// TIA Portal project "DATN" (V16)

(* hardware
DEVICE "S7-1200 station_1"  S7-1200 Station
   slot 0: "Rack_0"  S7-1200 Rack  Rack  V1.0
   slot 1: "PLC_1"  CPU 1214C DC/DC/DC  6ES7 214-1AG40-0XB0  V4.0
DEVICE "PC-System_1"  SIMATIC PC station
   slot 0: "SIMATIC PC station"  Rail  SIMATIC PC-Station  V1.0
      slot 125: "Stationmanager"  Station_Manager  V6.0.4
   slot 1: "HMI_RT_1"  WinCC RT Advanced  6AV2 104-0xxxx-xxxx  16.0.0.0
      slot 33792: "Computer interface"  Host interface
   slot 2: "IE general_1"  IE General  IE_CP  V8.2.0
*)

// ===== PLC "PLC_1"  CPU 1214C DC/DC/DC =====

VAR_GLOBAL   // PLC tag table "Default tag table"
   "System_Byte" AT %MB1000 : Byte;
   "FirstScan" AT %M1000.0 : Bool;
   "DiagStatusUpdate" AT %M1000.1 : Bool;
   "AlwaysTRUE" AT %M1000.2 : Bool;
   "AlwaysFALSE" AT %M1000.3 : Bool;
END_VAR

VAR_GLOBAL   // PLC tag table "1_IN"
   "CB_CAP_PHOI" AT %I0.0 : Bool;
   "CB_SP_1" AT %I0.1 : Bool;
   "CB_SP_2" AT %I0.2 : Bool;
   "CB_SP_3" AT %I0.3 : Bool;
   "PB_START" AT %I0.4 : Bool;
   "PB_STOP" AT %I0.5 : Bool;
   "PB_RESET" AT %I0.6 : Bool;
   "HMI_CB_CAP_PHOI" AT %M100.0 : Bool;
   "HMI_CB_SP_1" AT %M100.1 : Bool;
   "HMI_CB_SP_2" AT %M100.2 : Bool;
   "HMI_CB_SP_3" AT %M100.3 : Bool;
   "HMI_PB_START" AT %M100.4 : Bool;
   "HMI_PB_STOP" AT %M100.5 : Bool;
   "HMI_PB_RESET" AT %M100.6 : Bool;
   "MAN_BT" AT %M100.7 : Bool;
   "MAN_XYLANH_1" AT %M101.0 : Bool;
   "MAN_XYLANH_2" AT %M101.1 : Bool;
   "MAN_CAP_PHOI" AT %M101.2 : Bool;
   "HMI_AUTO_MAN" AT %M101.3 : Bool;
   "RST_SP_1" AT %M101.4 : Bool;
   "RST_SP_2" AT %M101.5 : Bool;
   "RST_SP_3" AT %M101.6 : Bool;
END_VAR

VAR_GLOBAL   // PLC tag table "2_OUT"
   "BANG_TAI" AT %Q0.0 : Bool;
   "XY_LANH_1" AT %Q0.1 : Bool;
   "XY_LANH_2" AT %Q0.2 : Bool;
   "DEN_START" AT %Q0.5 : Bool;
   "DEN_STOP" AT %Q0.6 : Bool;
   "XY_LANH_CAP_PHOI_1" AT %Q0.3 : Bool;
   "DEN_RESET" AT %Q0.7 : Bool;
END_VAR

VAR_GLOBAL   // PLC tag table "3_MEMORY"
   "SP_3" AT %M200.0 : Bool;
   "RUN_PHAN_LOAI" AT %M200.1 : Bool;
   "BT_1" AT %M200.2 : Bool;
   "BT_2" AT %M200.3 : Bool;
   "NGAT_CB_CAP_PHOI" AT %M200.4 : Bool;
   "RST_COUNTER_SP_1" AT %M200.5 : Bool;
   "RST_COUNTER_SP_2" AT %M200.6 : Bool;
   "RST_COUNTER_SP_3" AT %M200.7 : Bool;
   "den_rst_1" AT %M201.1 : Bool;
   "den_rst_2" AT %M201.2 : Bool;
   "NGAT_HE_THONG" AT %M201.3 : Bool;
   "OUT_counter_1" AT %M201.4 : Bool;
   "OUT_counter_2" AT %M201.5 : Bool;
   "OUT_counter_3" AT %M201.6 : Bool;
   "MODE_AUTO" AT %M201.7 : Bool;
   "MODE_MAN" AT %M202.0 : Bool;
   "xylanh_cap_phoi_auto" AT %M202.1 : Bool;
   "xylanh_cap_phoi_man" AT %M202.2 : Bool;
   "xylanh_1_auto" AT %M202.3 : Bool;
   "xylanh_1_man" AT %M202.4 : Bool;
   "xylanh_2_auto" AT %M202.5 : Bool;
   "xylanh_2_man" AT %M202.6 : Bool;
   "ngat_mau_sac" AT %M202.7 : Bool;
END_VAR

VAR_GLOBAL   // PLC tag table "5_M_TIME_500"
   "TIME_XY_LANH_1" AT %MD500 : Time;
   "TIME_XY_LANH_2" AT %MD504 : Time;
   "TIME_SP_3" AT %MD508 : Time;
   "TIME_CAP_PHOI" AT %MD512 : Time;
   "TIME_NGAT_CAP_PHOI" AT %MD516 : Time;
   "TIME_ERROR_KHONG_SP" AT %MD520 : Time;
   "TIME_ERROR_STUCK" AT %MD524 : Time;
END_VAR

VAR_GLOBAL   // PLC tag table "4_P_N_MEMORy"
   "N_CB_SP_1" AT %M300.0 : Bool;
   "N_CB_SP_2" AT %M300.1 : Bool;
   "N_CB_SP_3" AT %M300.2 : Bool;
   "N_XY_LANH_1" AT %M300.3 : Bool;
   "N_XY_LANH_2" AT %M300.4 : Bool;
   "N_SP_3" AT %M300.5 : Bool;
   "N_M_CB_SP_1" AT %M300.6 : Bool;
   "N_M_CB_SP_2" AT %M300.7 : Bool;
   "N_M_CB_SP_3" AT %M301.0 : Bool;
END_VAR

VAR_GLOBAL   // PLC tag table "6_DATA_real_int"
   "LUU_MAU" AT %MW222 : Int;
   "Mau Sac" AT %MW220 : Int;
END_VAR

VAR_GLOBAL   // PLC tag table "7_ALARM"
   "BIT_WARNING_KHONG_SP" AT %M400.0 : Bool;
   "DATA_WORD_WARNING" AT %MW400 : Int;
   "MULTI_ERROR" AT %M450.0 : Bool;
   "BIT_ERROR_STUCK_sp_1" AT %M402.0 : Bool;
   "BIT_ERROR_STUCK_sp_2" AT %M404.0 : Bool;
   "BIT_ERROR_STUCK_sp_3" AT %M406.0 : Bool;
   "DATA_WORD_ERROR_1" AT %MW402 : Int;
   "DATA_WORD_ERROR_2" AT %MW404 : Int;
   "DATA_WORD_ERROR_3" AT %MW406 : Int;
END_VAR

DATA_BLOCK "MB"   // DB12
{ S7_Optimized_Access := 'FALSE' }
VERSION : 0.1
   VAR
      DISCONNECT : Bool;
      H_reg : Array[0..10] of Int;
      CONNECT : TCON_IP_v4;
      ERROR : Bool;
      STATUS : Word;
   END_VAR
BEGIN
   CONNECT.InterfaceId := 64;
   CONNECT.ID := 1;
   CONNECT.ConnectionType := 11;
   CONNECT.ActiveEstablished := TRUE;
   CONNECT.RemoteAddress.ADDR[1] := 192;
   CONNECT.RemoteAddress.ADDR[2] := 168;
   CONNECT.RemoteAddress.ADDR[3] := 0;
   CONNECT.RemoteAddress.ADDR[4] := 10;
   CONNECT.LocalPort := 502;
   CONNECT.RemotePort := 0;
END_DATA_BLOCK

DATA_BLOCK "gh_sp"   // DB13
{ S7_Optimized_Access := 'TRUE' }
VERSION : 0.1
   VAR
      GH_SP_1 : USInt := 3;
      GH_SP_2 : USInt := 3;
      GH_SP_3 : USInt := 3;
   END_VAR
BEGIN
END_DATA_BLOCK

// folder: System blocks/Program resources

DATA_BLOCK "TIMER_CAP_PHOI"   // DB1
{ S7_Optimized_Access := 'TRUE' }
AUTHOR : Simatic
FAMILY : IEC
NAME : IEC_TMR
VERSION : 1.0
// stored: InstanceOfName IEC_TIMER
"IEC_TIMER"
BEGIN
END_DATA_BLOCK

DATA_BLOCK "TIMER_XY_LANH_1"   // DB2
{ S7_Optimized_Access := 'TRUE' }
AUTHOR : Simatic
FAMILY : IEC
NAME : IEC_TMR
VERSION : 1.0
// stored: InstanceOfName IEC_TIMER
"IEC_TIMER"
BEGIN
END_DATA_BLOCK

DATA_BLOCK "TIMER_XY_LANH_2"   // DB3
{ S7_Optimized_Access := 'TRUE' }
AUTHOR : Simatic
FAMILY : IEC
NAME : IEC_TMR
VERSION : 1.0
// stored: InstanceOfName IEC_TIMER
"IEC_TIMER"
BEGIN
END_DATA_BLOCK

DATA_BLOCK "TIMER_SP_3"   // DB4
{ S7_Optimized_Access := 'TRUE' }
AUTHOR : Simatic
FAMILY : IEC
NAME : IEC_TMR
VERSION : 1.0
// stored: InstanceOfName IEC_TIMER
"IEC_TIMER"
BEGIN
END_DATA_BLOCK

DATA_BLOCK "COUNTER_SP_1"   // DB5
{ S7_Optimized_Access := 'TRUE' }
AUTHOR : Simatic
FAMILY : IEC
NAME : CNTR
VERSION : 1.0
// stored: InstanceOfName IEC_COUNTER
"IEC_COUNTER"
BEGIN
END_DATA_BLOCK

DATA_BLOCK "COUNTER_SP_2"   // DB6
{ S7_Optimized_Access := 'TRUE' }
AUTHOR : Simatic
FAMILY : IEC
NAME : CNTR
VERSION : 1.0
// stored: InstanceOfName IEC_COUNTER
"IEC_COUNTER"
BEGIN
END_DATA_BLOCK

DATA_BLOCK "COUNTER_SP_3"   // DB7
{ S7_Optimized_Access := 'TRUE' }
AUTHOR : Simatic
FAMILY : IEC
NAME : CNTR
VERSION : 1.0
// stored: InstanceOfName IEC_COUNTER
"IEC_COUNTER"
BEGIN
END_DATA_BLOCK

DATA_BLOCK "TIMER_NGAT_CAP_PHOI"   // DB8
{ S7_Optimized_Access := 'TRUE' }
AUTHOR : Simatic
FAMILY : IEC
NAME : IEC_TMR
VERSION : 1.0
// stored: InstanceOfName IEC_TIMER
"IEC_TIMER"
BEGIN
END_DATA_BLOCK

DATA_BLOCK "TIMER_LOI_KHONG_SP"   // DB9
{ S7_Optimized_Access := 'TRUE' }
AUTHOR : Simatic
FAMILY : IEC
NAME : IEC_TMR
VERSION : 1.0
// stored: InstanceOfName IEC_TIMER
"IEC_TIMER"
BEGIN
END_DATA_BLOCK

DATA_BLOCK "TIMER_den_vang"   // DB10
{ S7_Optimized_Access := 'TRUE' }
AUTHOR : Simatic
FAMILY : IEC
NAME : IEC_TMR
VERSION : 1.0
// stored: InstanceOfName IEC_TIMER
"IEC_TIMER"
BEGIN
END_DATA_BLOCK

DATA_BLOCK "TIMER_STUCK_1"   // DB14
{ S7_Optimized_Access := 'TRUE' }
AUTHOR : Simatic
FAMILY : IEC
NAME : IEC_TMR
VERSION : 1.0
// stored: InstanceOfName IEC_TIMER
"IEC_TIMER"
BEGIN
END_DATA_BLOCK

DATA_BLOCK "TIMER_STUCK_2"   // DB15
{ S7_Optimized_Access := 'TRUE' }
AUTHOR : Simatic
FAMILY : IEC
NAME : IEC_TMR
VERSION : 1.0
// stored: InstanceOfName IEC_TIMER
"IEC_TIMER"
BEGIN
END_DATA_BLOCK

DATA_BLOCK "TIMER_STUCK_3"   // DB16
{ S7_Optimized_Access := 'TRUE' }
AUTHOR : Simatic
FAMILY : IEC
NAME : IEC_TMR
VERSION : 1.0
// stored: InstanceOfName IEC_TIMER
"IEC_TIMER"
BEGIN
END_DATA_BLOCK

// folder: (top level)

FUNCTION "FC_1_Modbus_TCP" : Void   // FC1, LAD
{ S7_Optimized_Access := 'TRUE' }
VERSION : 0.1
BEGIN

REGION Network 1
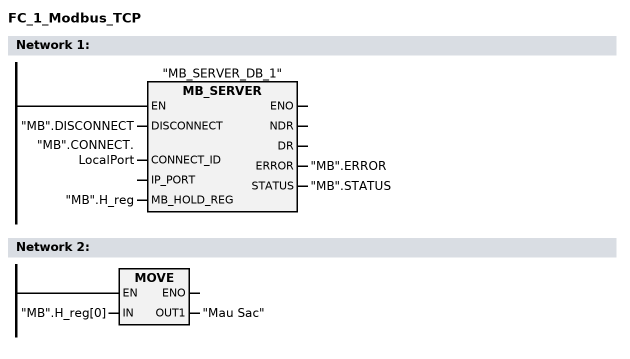
   "MB_SERVER_DB_1"(DISCONNECT := "MB".DISCONNECT,   // MB_SERVER
                    CONNECT_ID := "MB".CONNECT.LocalPort,
                    MB_HOLD_REG := "MB".H_reg,
                    ERROR => "MB".ERROR,
                    STATUS => "MB".STATUS);
END_REGION

REGION Network 2
   RUNG wire#powerrail
      Move(in := "MB".H_reg[0], out1 => "Mau Sac")
   END_RUNG
   // the same network as SCL:
   "Mau Sac" := "MB".H_reg[0];
END_REGION
END_FUNCTION

FUNCTION "FC_4_PHAN_LOAI_SP_1" : Void   // FC2, LAD
{ S7_Optimized_Access := 'TRUE' }
VERSION : 0.1
   VAR_TEMP   // added for the SCL form of the ladder/FBD networks
      _w1 : Bool;
      _w2 : Bool;
   END_VAR
BEGIN

REGION Network 1
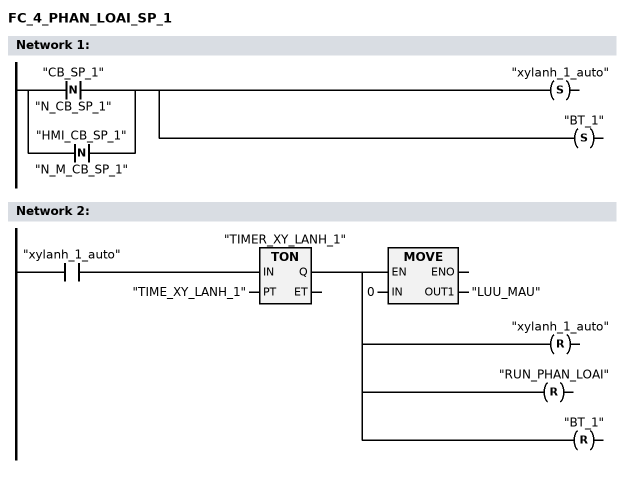
   RUNG wire#powerrail
      N_Contact(operand := "CB_SP_1", bit := "N_CB_SP_1")
      wire#w1
      S_Coil( "xylanh_1_auto" )
   END_RUNG
   RUNG wire#powerrail
      N_Contact(operand := "HMI_CB_SP_1", bit := "N_M_CB_SP_1")
   END_RUNG wire#w1
   RUNG wire#w1
      S_Coil( "BT_1" )
   END_RUNG
   // the same network as SCL:
   #_w1 := NOT "CB_SP_1" AND "N_CB_SP_1";   // falling edge of "CB_SP_1"
   "N_CB_SP_1" := "CB_SP_1";
   #_w2 := NOT "HMI_CB_SP_1" AND "N_M_CB_SP_1";   // falling edge of "HMI_CB_SP_1"
   "N_M_CB_SP_1" := "HMI_CB_SP_1";
   IF #_w1 OR #_w2 THEN
       "xylanh_1_auto" := TRUE;
       "BT_1" := TRUE;
   END_IF;
END_REGION

REGION Network 2
   "TIMER_XY_LANH_1".TON(IN := "xylanh_1_auto", PT := "TIME_XY_LANH_1");
   IF "TIMER_XY_LANH_1".Q THEN
       "LUU_MAU" := 0;
       "xylanh_1_auto" := FALSE;
       "RUN_PHAN_LOAI" := FALSE;
       "BT_1" := FALSE;
   END_IF;
END_REGION
END_FUNCTION

FUNCTION "FC_5_PHAN_LOAI_SP_2" : Void   // FC3, LAD
{ S7_Optimized_Access := 'TRUE' }
VERSION : 0.1
   VAR_TEMP   // added for the SCL form of the ladder/FBD networks
      _w1 : Bool;
      _w2 : Bool;
   END_VAR
BEGIN

REGION Network 1
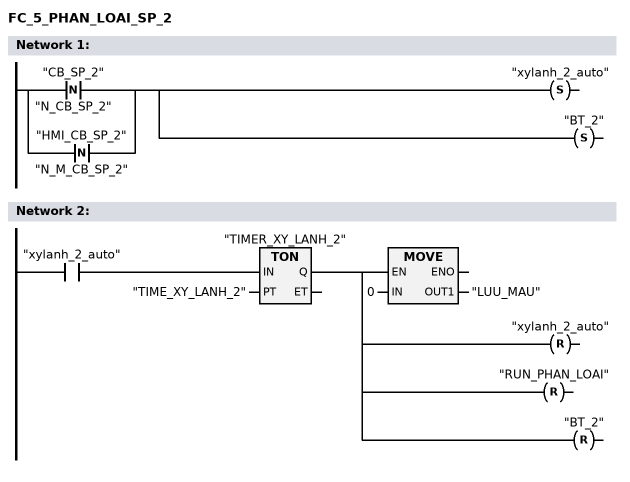
   RUNG wire#powerrail
      N_Contact(operand := "CB_SP_2", bit := "N_CB_SP_2")
      wire#w1
      S_Coil( "xylanh_2_auto" )
   END_RUNG
   RUNG wire#powerrail
      N_Contact(operand := "HMI_CB_SP_2", bit := "N_M_CB_SP_2")
   END_RUNG wire#w1
   RUNG wire#w1
      S_Coil( "BT_2" )
   END_RUNG
   // the same network as SCL:
   #_w1 := NOT "CB_SP_2" AND "N_CB_SP_2";   // falling edge of "CB_SP_2"
   "N_CB_SP_2" := "CB_SP_2";
   #_w2 := NOT "HMI_CB_SP_2" AND "N_M_CB_SP_2";   // falling edge of "HMI_CB_SP_2"
   "N_M_CB_SP_2" := "HMI_CB_SP_2";
   IF #_w1 OR #_w2 THEN
       "xylanh_2_auto" := TRUE;
       "BT_2" := TRUE;
   END_IF;
END_REGION

REGION Network 2
   "TIMER_XY_LANH_2".TON(IN := "xylanh_2_auto", PT := "TIME_XY_LANH_2");
   IF "TIMER_XY_LANH_2".Q THEN
       "LUU_MAU" := 0;
       "xylanh_2_auto" := FALSE;
       "RUN_PHAN_LOAI" := FALSE;
       "BT_2" := FALSE;
   END_IF;
END_REGION
END_FUNCTION

FUNCTION "FC_6_PHAN_LOAI_SP_3" : Void   // FC4, LAD
{ S7_Optimized_Access := 'TRUE' }
VERSION : 0.1
   VAR_TEMP   // added for the SCL form of the ladder/FBD networks
      _w1 : Bool;
      _w2 : Bool;
   END_VAR
BEGIN

REGION Network 1
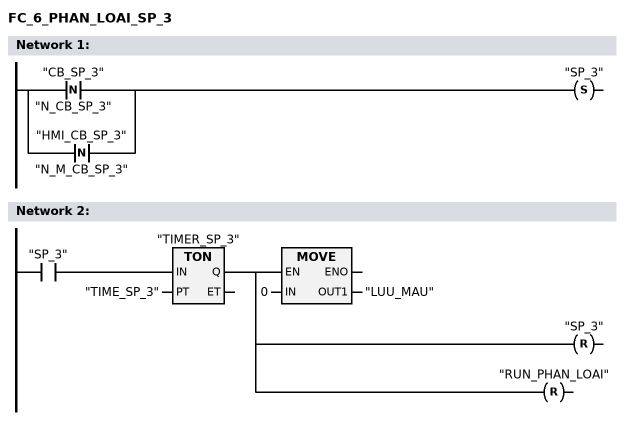
   RUNG wire#powerrail
      N_Contact(operand := "CB_SP_3", bit := "N_CB_SP_3")
      wire#w1
      S_Coil( "SP_3" )
   END_RUNG
   RUNG wire#powerrail
      N_Contact(operand := "HMI_CB_SP_3", bit := "N_M_CB_SP_3")
   END_RUNG wire#w1
   // the same network as SCL:
   #_w1 := NOT "CB_SP_3" AND "N_CB_SP_3";   // falling edge of "CB_SP_3"
   "N_CB_SP_3" := "CB_SP_3";
   #_w2 := NOT "HMI_CB_SP_3" AND "N_M_CB_SP_3";   // falling edge of "HMI_CB_SP_3"
   "N_M_CB_SP_3" := "HMI_CB_SP_3";
   IF #_w1 OR #_w2 THEN "SP_3" := TRUE; END_IF;
END_REGION

REGION Network 2
   "TIMER_SP_3".TON(IN := "SP_3", PT := "TIME_SP_3");
   IF "TIMER_SP_3".Q THEN
       "LUU_MAU" := 0;
       "SP_3" := FALSE;
       "RUN_PHAN_LOAI" := FALSE;
   END_IF;
END_REGION
END_FUNCTION

FUNCTION "FC_3_CAP_PHOI_TU_DONG" : Void   // FC5, LAD
{ S7_Optimized_Access := 'TRUE' }
VERSION : 0.1
BEGIN

REGION Network 1
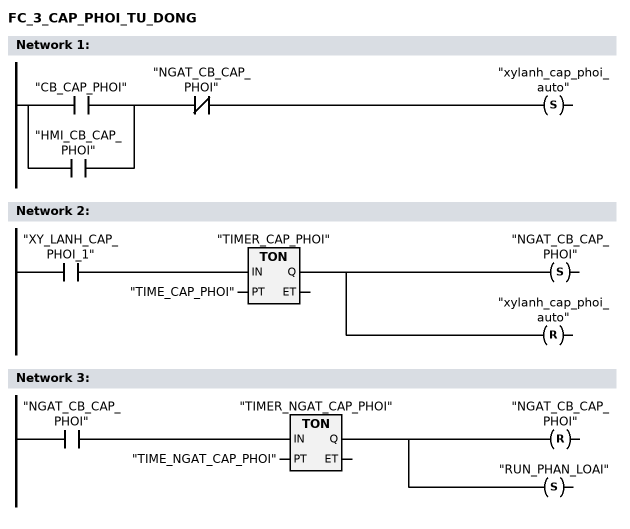
   RUNG wire#powerrail
      Contact( "CB_CAP_PHOI" )
      wire#w1
      I_Contact( "NGAT_CB_CAP_PHOI" )
      S_Coil( "xylanh_cap_phoi_auto" )
   END_RUNG
   RUNG wire#powerrail
      Contact( "HMI_CB_CAP_PHOI" )
   END_RUNG wire#w1
   // the same network as SCL:
   IF ("CB_CAP_PHOI" OR "HMI_CB_CAP_PHOI") AND NOT "NGAT_CB_CAP_PHOI" THEN
       "xylanh_cap_phoi_auto" := TRUE;
   END_IF;
END_REGION

REGION Network 2
   "TIMER_CAP_PHOI".TON(IN := "XY_LANH_CAP_PHOI_1", PT := "TIME_CAP_PHOI");
   IF "TIMER_CAP_PHOI".Q THEN
       "NGAT_CB_CAP_PHOI" := TRUE;
       "xylanh_cap_phoi_auto" := FALSE;
   END_IF;
END_REGION

REGION Network 3
   "TIMER_NGAT_CAP_PHOI".TON(IN := "NGAT_CB_CAP_PHOI", PT := "TIME_NGAT_CAP_PHOI");
   IF "TIMER_NGAT_CAP_PHOI".Q THEN
       "NGAT_CB_CAP_PHOI" := FALSE;
       "RUN_PHAN_LOAI" := TRUE;
   END_IF;
END_REGION
END_FUNCTION

FUNCTION "FC_2_RESET_HE_THONG" : Void   // FC6, LAD
{ S7_Optimized_Access := 'TRUE' }
VERSION : 0.1
BEGIN

REGION Network 1
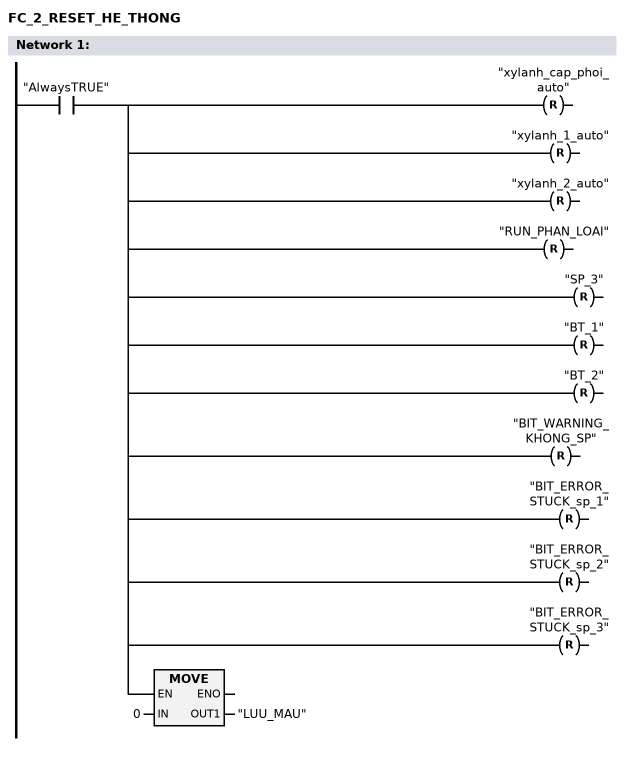
   RUNG wire#powerrail
      Contact( "AlwaysTRUE" )
      wire#w1
      R_Coil( "xylanh_cap_phoi_auto" )
   END_RUNG
   RUNG wire#w1
      R_Coil( "xylanh_1_auto" )
   END_RUNG
   RUNG wire#w1
      R_Coil( "xylanh_2_auto" )
   END_RUNG
   RUNG wire#w1
      R_Coil( "RUN_PHAN_LOAI" )
   END_RUNG
   RUNG wire#w1
      R_Coil( "SP_3" )
   END_RUNG
   RUNG wire#w1
      R_Coil( "BT_1" )
   END_RUNG
   RUNG wire#w1
      R_Coil( "BT_2" )
   END_RUNG
   RUNG wire#w1
      R_Coil( "BIT_WARNING_KHONG_SP" )
   END_RUNG
   RUNG wire#w1
      R_Coil( "BIT_ERROR_STUCK_sp_1" )
   END_RUNG
   RUNG wire#w1
      R_Coil( "BIT_ERROR_STUCK_sp_2" )
   END_RUNG
   RUNG wire#w1
      R_Coil( "BIT_ERROR_STUCK_sp_3" )
   END_RUNG
   RUNG wire#w1
      Move(in := 0, out1 => "LUU_MAU")
   END_RUNG
   // the same network as SCL:
   IF "AlwaysTRUE" THEN
       "xylanh_cap_phoi_auto" := FALSE;
       "xylanh_1_auto" := FALSE;
       "xylanh_2_auto" := FALSE;
       "RUN_PHAN_LOAI" := FALSE;
       "SP_3" := FALSE;
       "BT_1" := FALSE;
       "BT_2" := FALSE;
       "BIT_WARNING_KHONG_SP" := FALSE;
       "BIT_ERROR_STUCK_sp_1" := FALSE;
       "BIT_ERROR_STUCK_sp_2" := FALSE;
       "BIT_ERROR_STUCK_sp_3" := FALSE;
       "LUU_MAU" := 0;
   END_IF;
END_REGION
END_FUNCTION

FUNCTION "FC_7_COUNTER_SP" : Void   // FC7, LAD
{ S7_Optimized_Access := 'TRUE' }
VERSION : 0.1
   VAR_TEMP   // added for the SCL form of the ladder/FBD networks
      _w1 : Bool;
   END_VAR
BEGIN

REGION Network 1
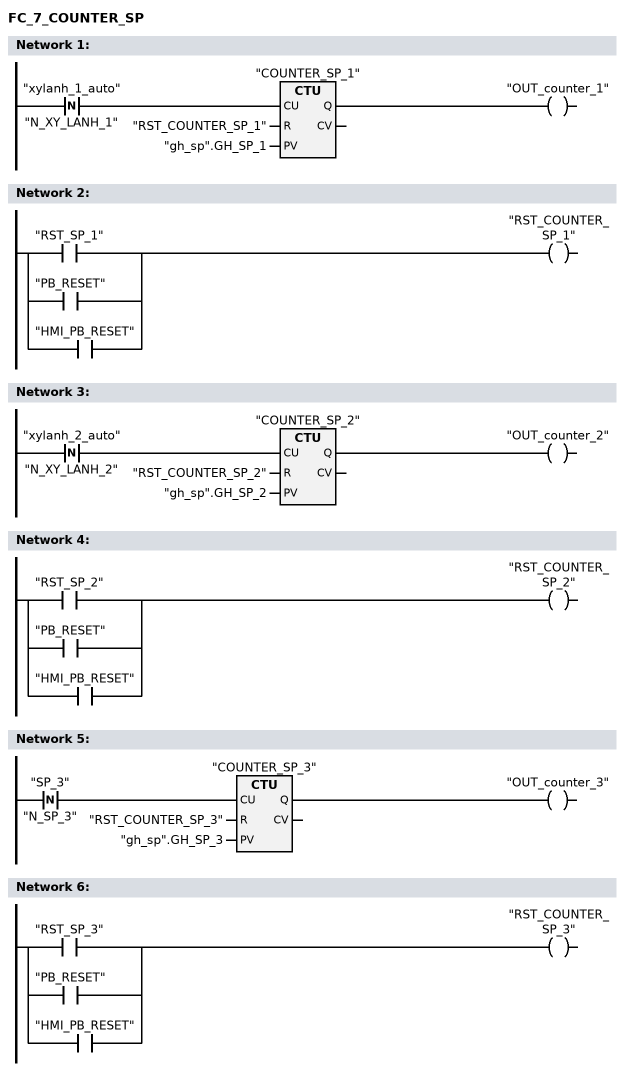
   #_w1 := NOT "xylanh_1_auto" AND "N_XY_LANH_1";   // falling edge of "xylanh_1_auto"
   "N_XY_LANH_1" := "xylanh_1_auto";
   "COUNTER_SP_1".CTU(CU := #_w1, R := "RST_COUNTER_SP_1", PV := "gh_sp".GH_SP_1);
   "OUT_counter_1" := "COUNTER_SP_1".Q;
END_REGION

REGION Network 2
   RUNG wire#powerrail
      Contact( "RST_SP_1" )
      wire#w1
      Coil( "RST_COUNTER_SP_1" )
   END_RUNG
   RUNG wire#powerrail
      Contact( "PB_RESET" )
   END_RUNG wire#w1
   RUNG wire#powerrail
      Contact( "HMI_PB_RESET" )
   END_RUNG wire#w1
   // the same network as SCL:
   "RST_COUNTER_SP_1" := "RST_SP_1" OR "PB_RESET" OR "HMI_PB_RESET";
END_REGION

REGION Network 3
   #_w1 := NOT "xylanh_2_auto" AND "N_XY_LANH_2";   // falling edge of "xylanh_2_auto"
   "N_XY_LANH_2" := "xylanh_2_auto";
   "COUNTER_SP_2".CTU(CU := #_w1, R := "RST_COUNTER_SP_2", PV := "gh_sp".GH_SP_2);
   "OUT_counter_2" := "COUNTER_SP_2".Q;
END_REGION

REGION Network 4
   RUNG wire#powerrail
      Contact( "RST_SP_2" )
      wire#w1
      Coil( "RST_COUNTER_SP_2" )
   END_RUNG
   RUNG wire#powerrail
      Contact( "PB_RESET" )
   END_RUNG wire#w1
   RUNG wire#powerrail
      Contact( "HMI_PB_RESET" )
   END_RUNG wire#w1
   // the same network as SCL:
   "RST_COUNTER_SP_2" := "RST_SP_2" OR "PB_RESET" OR "HMI_PB_RESET";
END_REGION

REGION Network 5
   #_w1 := NOT "SP_3" AND "N_SP_3";   // falling edge of "SP_3"
   "N_SP_3" := "SP_3";
   "COUNTER_SP_3".CTU(CU := #_w1, R := "RST_COUNTER_SP_3", PV := "gh_sp".GH_SP_3);
   "OUT_counter_3" := "COUNTER_SP_3".Q;
END_REGION

REGION Network 6
   RUNG wire#powerrail
      Contact( "RST_SP_3" )
      wire#w1
      Coil( "RST_COUNTER_SP_3" )
   END_RUNG
   RUNG wire#powerrail
      Contact( "PB_RESET" )
   END_RUNG wire#w1
   RUNG wire#powerrail
      Contact( "HMI_PB_RESET" )
   END_RUNG wire#w1
   // the same network as SCL:
   "RST_COUNTER_SP_3" := "RST_SP_3" OR "PB_RESET" OR "HMI_PB_RESET";
END_REGION
END_FUNCTION

FUNCTION "FC_8_ERROR_KHONG_SP" : Void   // FC8, LAD
{ S7_Optimized_Access := 'TRUE' }
VERSION : 0.1
BEGIN

REGION Network 1
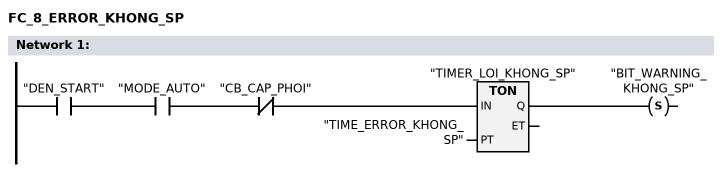
   "TIMER_LOI_KHONG_SP".TON(IN := "DEN_START" AND "MODE_AUTO" AND NOT "CB_CAP_PHOI",
                           PT := "TIME_ERROR_KHONG_SP");
   IF "TIMER_LOI_KHONG_SP".Q THEN "BIT_WARNING_KHONG_SP" := TRUE; END_IF;
END_REGION
END_FUNCTION

FUNCTION "FC_9_ERROR_STUCK" : Void   // FC9, LAD
{ S7_Optimized_Access := 'TRUE' }
VERSION : 0.1
BEGIN

REGION Network 1
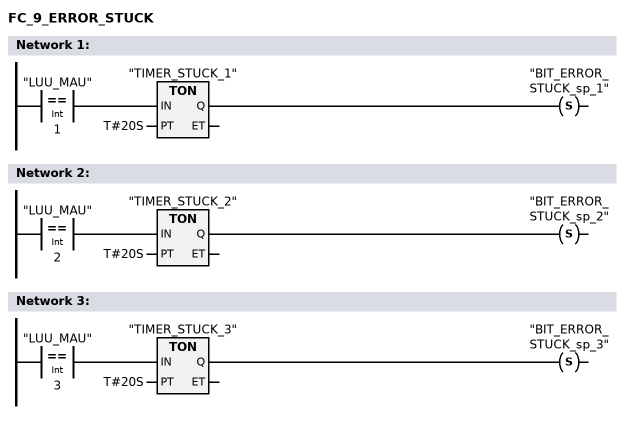
   "TIMER_STUCK_1".TON(IN := "LUU_MAU" = 1, PT := T#20S);
   IF "TIMER_STUCK_1".Q THEN "BIT_ERROR_STUCK_sp_1" := TRUE; END_IF;
END_REGION

REGION Network 2
   "TIMER_STUCK_2".TON(IN := "LUU_MAU" = 2, PT := T#20S);
   IF "TIMER_STUCK_2".Q THEN "BIT_ERROR_STUCK_sp_2" := TRUE; END_IF;
END_REGION

REGION Network 3
   "TIMER_STUCK_3".TON(IN := "LUU_MAU" = 3, PT := T#20S);
   IF "TIMER_STUCK_3".Q THEN "BIT_ERROR_STUCK_sp_3" := TRUE; END_IF;
END_REGION
END_FUNCTION

FUNCTION "FC_10_multierror" : Void   // FC10, LAD
{ S7_Optimized_Access := 'TRUE' }
VERSION : 0.1
BEGIN

REGION Network 1
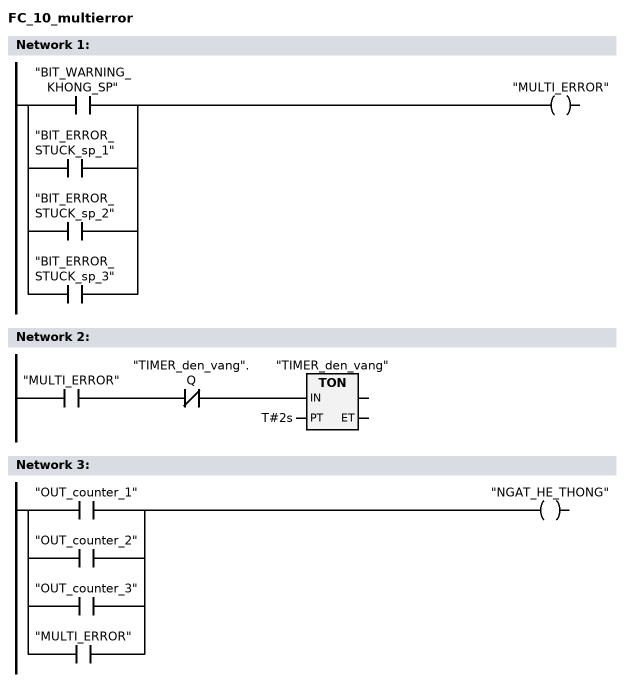
   RUNG wire#powerrail
      Contact( "BIT_WARNING_KHONG_SP" )
      wire#w1
      Coil( "MULTI_ERROR" )
   END_RUNG
   RUNG wire#powerrail
      Contact( "BIT_ERROR_STUCK_sp_1" )
   END_RUNG wire#w1
   RUNG wire#powerrail
      Contact( "BIT_ERROR_STUCK_sp_2" )
   END_RUNG wire#w1
   RUNG wire#powerrail
      Contact( "BIT_ERROR_STUCK_sp_3" )
   END_RUNG wire#w1
   // the same network as SCL:
   "MULTI_ERROR" := "BIT_WARNING_KHONG_SP" OR "BIT_ERROR_STUCK_sp_1" OR "BIT_ERROR_STUCK_sp_2" OR "BIT_ERROR_STUCK_sp_3";
END_REGION

REGION Network 2
   "TIMER_den_vang".TON(IN := "MULTI_ERROR" AND NOT "TIMER_den_vang".Q, PT := T#2s);
END_REGION

REGION Network 3
   RUNG wire#powerrail
      Contact( "OUT_counter_1" )
      wire#w1
      Coil( "NGAT_HE_THONG" )
   END_RUNG
   RUNG wire#powerrail
      Contact( "OUT_counter_2" )
   END_RUNG wire#w1
   RUNG wire#powerrail
      Contact( "OUT_counter_3" )
   END_RUNG wire#w1
   RUNG wire#powerrail
      Contact( "MULTI_ERROR" )
   END_RUNG wire#w1
   // the same network as SCL:
   "NGAT_HE_THONG" := "OUT_counter_1" OR "OUT_counter_2" OR "OUT_counter_3" OR "MULTI_ERROR";
END_REGION
END_FUNCTION

ORGANIZATION_BLOCK "Main"   // OB1, LAD, ProgramCycle
TITLE = "Main Program Sweep (Cycle)"
{ S7_Optimized_Access := 'TRUE' }
VERSION : 0.1
   VAR_INPUT
      Initial_Call : Bool;   // Initial call of this OB
      Remanence : Bool;   // =True, if remanent data are available
   END_VAR
   VAR_TEMP
      Barcode_HMI : DWord;
   END_VAR
   VAR_TEMP   // added for the SCL form of the ladder/FBD networks
      _w1 : Bool;
   END_VAR
BEGIN

REGION Network 1
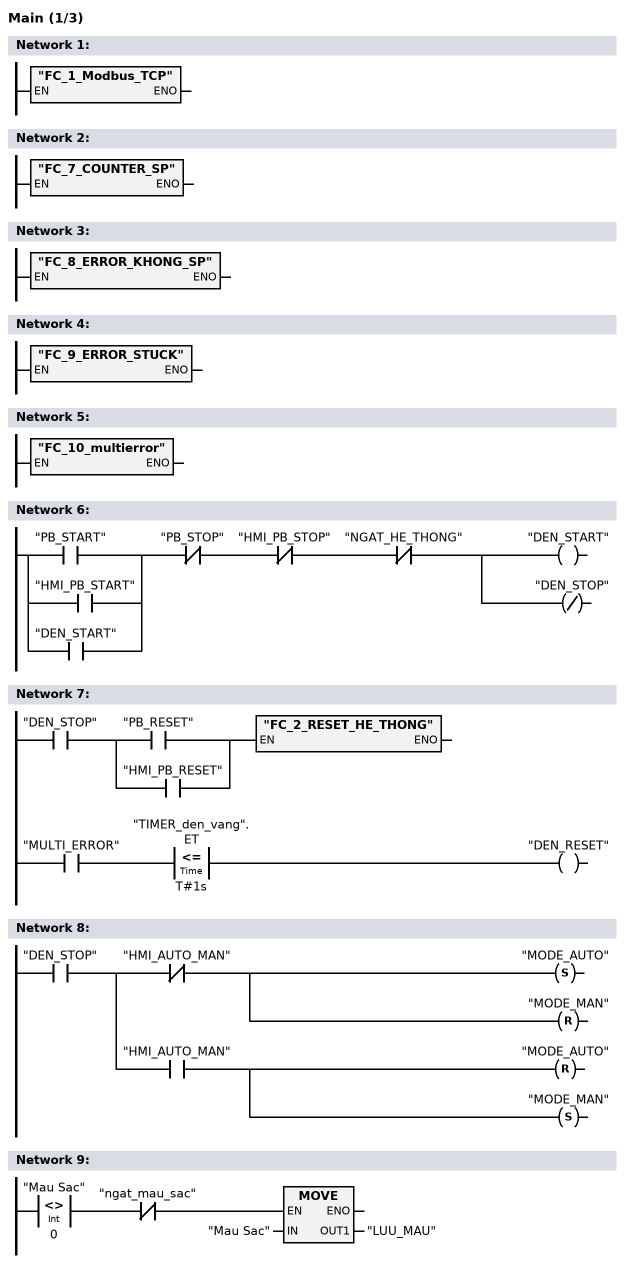
   RUNG wire#powerrail
      "FC_1_Modbus_TCP"()
   END_RUNG
   // the same network as SCL:
   "FC_1_Modbus_TCP"();
END_REGION

REGION Network 2
   RUNG wire#powerrail
      "FC_7_COUNTER_SP"()
   END_RUNG
   // the same network as SCL:
   "FC_7_COUNTER_SP"();
END_REGION

REGION Network 3
   RUNG wire#powerrail
      "FC_8_ERROR_KHONG_SP"()
   END_RUNG
   // the same network as SCL:
   "FC_8_ERROR_KHONG_SP"();
END_REGION

REGION Network 4
   RUNG wire#powerrail
      "FC_9_ERROR_STUCK"()
   END_RUNG
   // the same network as SCL:
   "FC_9_ERROR_STUCK"();
END_REGION

REGION Network 5
   RUNG wire#powerrail
      "FC_10_multierror"()
   END_RUNG
   // the same network as SCL:
   "FC_10_multierror"();
END_REGION

REGION Network 6
   RUNG wire#powerrail
      Contact( "PB_START" )
      wire#w1
      I_Contact( "PB_STOP" )
      I_Contact( "HMI_PB_STOP" )
      I_Contact( "NGAT_HE_THONG" )
      wire#w2
      Coil( "DEN_START" )
   END_RUNG
   RUNG wire#powerrail
      Contact( "HMI_PB_START" )
   END_RUNG wire#w1
   RUNG wire#powerrail
      Contact( "DEN_START" )
   END_RUNG wire#w1
   RUNG wire#w2
      I_Coil( "DEN_STOP" )
   END_RUNG
   // the same network as SCL:
   "DEN_START" := ("PB_START" OR "HMI_PB_START" OR "DEN_START") AND NOT "PB_STOP" AND NOT "HMI_PB_STOP" AND NOT "NGAT_HE_THONG";
   "DEN_STOP" := NOT "DEN_START";
END_REGION

REGION Network 7
   RUNG wire#powerrail
      Contact( "DEN_STOP" )
      wire#w1
      Contact( "PB_RESET" )
      wire#w2
      "FC_2_RESET_HE_THONG"()
   END_RUNG
   RUNG wire#w1
      Contact( "HMI_PB_RESET" )
   END_RUNG wire#w2
   RUNG wire#powerrail
      Contact( "MULTI_ERROR" )
      { S7_Templates := "SrcType := Time" } LE_Contact(in1 := "TIMER_den_vang".ET, in2 := T#1s)
      Coil( "DEN_RESET" )
   END_RUNG
   // the same network as SCL:
   IF "DEN_STOP" AND ("PB_RESET" OR "HMI_PB_RESET") THEN "FC_2_RESET_HE_THONG"(); END_IF;
   "DEN_RESET" := "MULTI_ERROR" AND ("TIMER_den_vang".ET <= T#1s);
END_REGION

REGION Network 8
   RUNG wire#powerrail
      Contact( "DEN_STOP" )
      wire#w1
      I_Contact( "HMI_AUTO_MAN" )
      wire#w2
      S_Coil( "MODE_AUTO" )
   END_RUNG
   RUNG wire#w2
      R_Coil( "MODE_MAN" )
   END_RUNG
   RUNG wire#w1
      Contact( "HMI_AUTO_MAN" )
      wire#w3
      R_Coil( "MODE_AUTO" )
   END_RUNG
   RUNG wire#w3
      S_Coil( "MODE_MAN" )
   END_RUNG
   // the same network as SCL:
   IF "DEN_STOP" AND NOT "HMI_AUTO_MAN" THEN
       "MODE_AUTO" := TRUE;
       "MODE_MAN" := FALSE;
   END_IF;
   IF "DEN_STOP" AND "HMI_AUTO_MAN" THEN
       "MODE_AUTO" := FALSE;
       "MODE_MAN" := TRUE;
   END_IF;
END_REGION

REGION Network 9
   RUNG wire#powerrail
      { S7_Templates := "SrcType := Int" } NE_Contact(in1 := "Mau Sac", in2 := 0)
      I_Contact( "ngat_mau_sac" )
      Move(in := "Mau Sac", out1 => "LUU_MAU")
   END_RUNG
   // the same network as SCL:
   IF ("Mau Sac" <> 0) AND NOT "ngat_mau_sac" THEN "LUU_MAU" := "Mau Sac"; END_IF;
END_REGION

REGION Network 10
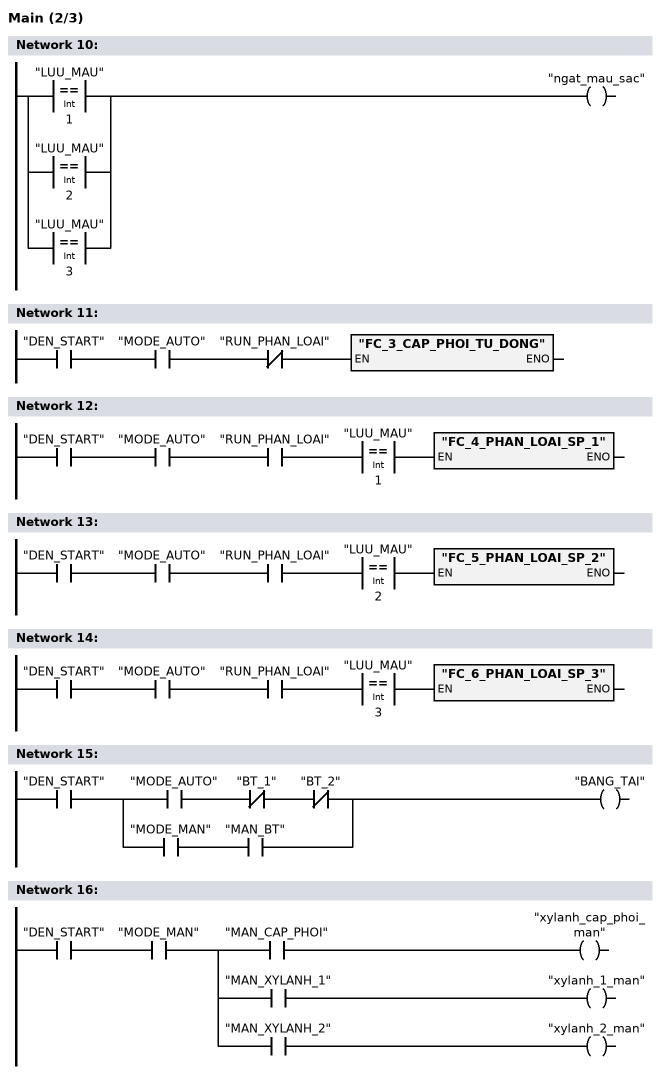
   RUNG wire#powerrail
      { S7_Templates := "SrcType := Int" } EQ_Contact(in1 := "LUU_MAU", in2 := 1)
      wire#w1
      Coil( "ngat_mau_sac" )
   END_RUNG
   RUNG wire#powerrail
      { S7_Templates := "SrcType := Int" } EQ_Contact(in1 := "LUU_MAU", in2 := 2)
   END_RUNG wire#w1
   RUNG wire#powerrail
      { S7_Templates := "SrcType := Int" } EQ_Contact(in1 := "LUU_MAU", in2 := 3)
   END_RUNG wire#w1
   // the same network as SCL:
   "ngat_mau_sac" := ("LUU_MAU" = 1) OR ("LUU_MAU" = 2) OR ("LUU_MAU" = 3);
END_REGION

REGION Network 11
   RUNG wire#powerrail
      Contact( "DEN_START" )
      Contact( "MODE_AUTO" )
      I_Contact( "RUN_PHAN_LOAI" )
      "FC_3_CAP_PHOI_TU_DONG"()
   END_RUNG
   // the same network as SCL:
   IF "DEN_START" AND "MODE_AUTO" AND NOT "RUN_PHAN_LOAI" THEN "FC_3_CAP_PHOI_TU_DONG"(); END_IF;
END_REGION

REGION Network 12
   RUNG wire#powerrail
      Contact( "DEN_START" )
      Contact( "MODE_AUTO" )
      Contact( "RUN_PHAN_LOAI" )
      { S7_Templates := "SrcType := Int" } EQ_Contact(in1 := "LUU_MAU", in2 := 1)
      "FC_4_PHAN_LOAI_SP_1"()
   END_RUNG
   // the same network as SCL:
   IF "DEN_START" AND "MODE_AUTO" AND "RUN_PHAN_LOAI" AND ("LUU_MAU" = 1) THEN
       "FC_4_PHAN_LOAI_SP_1"();
   END_IF;
END_REGION

REGION Network 13
   RUNG wire#powerrail
      Contact( "DEN_START" )
      Contact( "MODE_AUTO" )
      Contact( "RUN_PHAN_LOAI" )
      { S7_Templates := "SrcType := Int" } EQ_Contact(in1 := "LUU_MAU", in2 := 2)
      "FC_5_PHAN_LOAI_SP_2"()
   END_RUNG
   // the same network as SCL:
   IF "DEN_START" AND "MODE_AUTO" AND "RUN_PHAN_LOAI" AND ("LUU_MAU" = 2) THEN
       "FC_5_PHAN_LOAI_SP_2"();
   END_IF;
END_REGION

REGION Network 14
   RUNG wire#powerrail
      Contact( "DEN_START" )
      Contact( "MODE_AUTO" )
      Contact( "RUN_PHAN_LOAI" )
      { S7_Templates := "SrcType := Int" } EQ_Contact(in1 := "LUU_MAU", in2 := 3)
      "FC_6_PHAN_LOAI_SP_3"()
   END_RUNG
   // the same network as SCL:
   IF "DEN_START" AND "MODE_AUTO" AND "RUN_PHAN_LOAI" AND ("LUU_MAU" = 3) THEN
       "FC_6_PHAN_LOAI_SP_3"();
   END_IF;
END_REGION

REGION Network 15
   RUNG wire#powerrail
      Contact( "DEN_START" )
      wire#w1
      Contact( "MODE_AUTO" )
      I_Contact( "BT_1" )
      I_Contact( "BT_2" )
      wire#w2
      Coil( "BANG_TAI" )
   END_RUNG
   RUNG wire#w1
      Contact( "MODE_MAN" )
      Contact( "MAN_BT" )
   END_RUNG wire#w2
   // the same network as SCL:
   "BANG_TAI" := "DEN_START" AND (("MODE_AUTO" AND NOT "BT_1" AND NOT "BT_2") OR ("MODE_MAN" AND "MAN_BT"));
END_REGION

REGION Network 16
   RUNG wire#powerrail
      Contact( "DEN_START" )
      Contact( "MODE_MAN" )
      wire#w1
      Contact( "MAN_CAP_PHOI" )
      Coil( "xylanh_cap_phoi_man" )
   END_RUNG
   RUNG wire#w1
      Contact( "MAN_XYLANH_1" )
      Coil( "xylanh_1_man" )
   END_RUNG
   RUNG wire#w1
      Contact( "MAN_XYLANH_2" )
      Coil( "xylanh_2_man" )
   END_RUNG
   // the same network as SCL:
   #_w1 := "DEN_START" AND "MODE_MAN";
   "xylanh_cap_phoi_man" := #_w1 AND "MAN_CAP_PHOI";
   "xylanh_1_man" := #_w1 AND "MAN_XYLANH_1";
   "xylanh_2_man" := #_w1 AND "MAN_XYLANH_2";
END_REGION

REGION Network 17
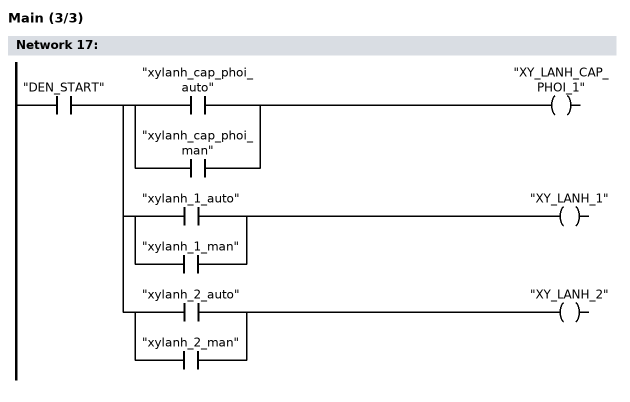
   RUNG wire#powerrail
      Contact( "DEN_START" )
      wire#w1
      Contact( "xylanh_cap_phoi_auto" )
      wire#w2
      Coil( "XY_LANH_CAP_PHOI_1" )
   END_RUNG
   RUNG wire#w1
      Contact( "xylanh_cap_phoi_man" )
   END_RUNG wire#w2
   RUNG wire#w1
      Contact( "xylanh_1_auto" )
      wire#w3
      Coil( "XY_LANH_1" )
   END_RUNG
   RUNG wire#w1
      Contact( "xylanh_1_man" )
   END_RUNG wire#w3
   RUNG wire#w1
      Contact( "xylanh_2_auto" )
      wire#w4
      Coil( "XY_LANH_2" )
   END_RUNG
   RUNG wire#w1
      Contact( "xylanh_2_man" )
   END_RUNG wire#w4
   // the same network as SCL:
   "XY_LANH_CAP_PHOI_1" := "DEN_START" AND ("xylanh_cap_phoi_auto" OR "xylanh_cap_phoi_man");
   "XY_LANH_1" := "DEN_START" AND ("xylanh_1_auto" OR "xylanh_1_man");
   "XY_LANH_2" := "DEN_START" AND ("xylanh_2_auto" OR "xylanh_2_man");
END_REGION
END_ORGANIZATION_BLOCK

ORGANIZATION_BLOCK "Startup"   // OB100, LAD, Startup
TITLE = "Complete Restart"
{ S7_Optimized_Access := 'TRUE' }
VERSION : 0.1
   VAR_INPUT
      LostRetentive : Bool;   // True if retentive data are lost
      LostRTC : Bool;   // True if date and time are lost
   END_VAR
BEGIN

REGION Network 1